FUNCTION "SEQUENCE_TRANSFER" : Void   // FC9, LAD
{ S7_Optimized_Access := 'TRUE' }
VERSION : 0.1
   VAR_TEMP   // added for the SCL form of the ladder/FBD networks
      _w1 : Bool;
      _w2 : Bool;
      _w3 : Bool;
      _w4 : Bool;
      _w5 : Bool;
      _w6 : Bool;
      _w7 : Bool;
      _w8 : Bool;
      _w9 : Bool;
      _w10 : Bool;
      _w11 : Bool;
      _w12 : Bool;
      _w13 : Bool;
      _w14 : Bool;
      _w15 : Bool;
      _w16 : Bool;
      _w17 : Bool;
      _w18 : Bool;
      _s5time1 : S5Time;
      _s5time2 : S5Time;
   END_VAR
BEGIN

REGION Network 1: START TRANSFER
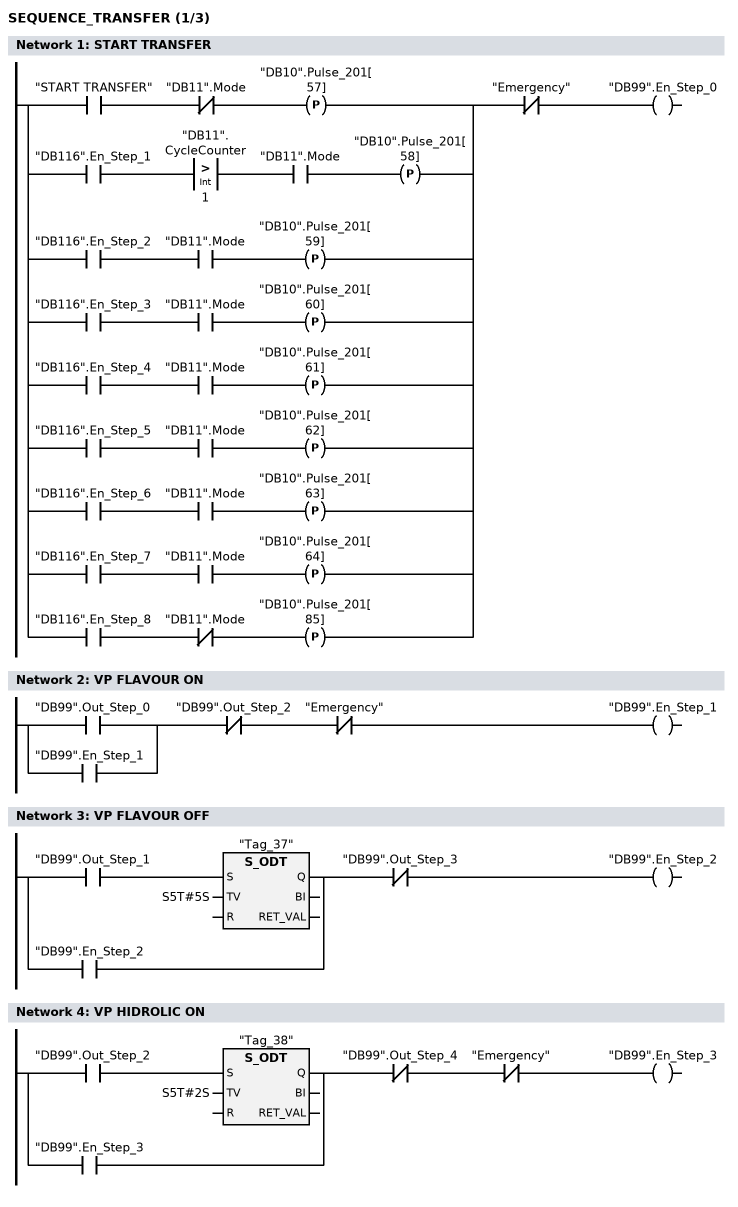
   RUNG wire#powerrail
      Contact( "START TRANSFER" )
      I_Contact( "DB11".Mode )
      P_Trig( "DB10".Pulse_201[57] )
      wire#w1
      I_Contact( "Emergency" )
      Coil( "DB99".En_Step_0 )
   END_RUNG
   RUNG wire#powerrail
      Contact( "DB116".En_Step_1 )
      { S7_Templates := "SrcType := Int" } GT_Contact(in1 := "DB11".CycleCounter, in2 := 1)
      Contact( "DB11".Mode )
      P_Trig( "DB10".Pulse_201[58] )
   END_RUNG wire#w1
   RUNG wire#powerrail
      Contact( "DB116".En_Step_2 )
      Contact( "DB11".Mode )
      P_Trig( "DB10".Pulse_201[59] )
   END_RUNG wire#w1
   RUNG wire#powerrail
      Contact( "DB116".En_Step_3 )
      Contact( "DB11".Mode )
      P_Trig( "DB10".Pulse_201[60] )
   END_RUNG wire#w1
   RUNG wire#powerrail
      Contact( "DB116".En_Step_4 )
      Contact( "DB11".Mode )
      P_Trig( "DB10".Pulse_201[61] )
   END_RUNG wire#w1
   RUNG wire#powerrail
      Contact( "DB116".En_Step_5 )
      Contact( "DB11".Mode )
      P_Trig( "DB10".Pulse_201[62] )
   END_RUNG wire#w1
   RUNG wire#powerrail
      Contact( "DB116".En_Step_6 )
      Contact( "DB11".Mode )
      P_Trig( "DB10".Pulse_201[63] )
   END_RUNG wire#w1
   RUNG wire#powerrail
      Contact( "DB116".En_Step_7 )
      Contact( "DB11".Mode )
      P_Trig( "DB10".Pulse_201[64] )
   END_RUNG wire#w1
   RUNG wire#powerrail
      Contact( "DB116".En_Step_8 )
      I_Contact( "DB11".Mode )
      P_Trig( "DB10".Pulse_201[85] )
   END_RUNG wire#w1
   // the same network as SCL:
   #_w1 := "START TRANSFER" AND NOT "DB11".Mode;
   #_w2 := #_w1 AND NOT "DB10".Pulse_201[57];   // rising edge
   "DB10".Pulse_201[57] := #_w1;
   #_w3 := "DB116".En_Step_1 AND ("DB11".CycleCounter > 1) AND "DB11".Mode;
   #_w4 := #_w3 AND NOT "DB10".Pulse_201[58];   // rising edge
   "DB10".Pulse_201[58] := #_w3;
   #_w5 := "DB116".En_Step_2 AND "DB11".Mode;
   #_w6 := #_w5 AND NOT "DB10".Pulse_201[59];   // rising edge
   "DB10".Pulse_201[59] := #_w5;
   #_w7 := "DB116".En_Step_3 AND "DB11".Mode;
   #_w8 := #_w7 AND NOT "DB10".Pulse_201[60];   // rising edge
   "DB10".Pulse_201[60] := #_w7;
   #_w9 := "DB116".En_Step_4 AND "DB11".Mode;
   #_w10 := #_w9 AND NOT "DB10".Pulse_201[61];   // rising edge
   "DB10".Pulse_201[61] := #_w9;
   #_w11 := "DB116".En_Step_5 AND "DB11".Mode;
   #_w12 := #_w11 AND NOT "DB10".Pulse_201[62];   // rising edge
   "DB10".Pulse_201[62] := #_w11;
   #_w13 := "DB116".En_Step_6 AND "DB11".Mode;
   #_w14 := #_w13 AND NOT "DB10".Pulse_201[63];   // rising edge
   "DB10".Pulse_201[63] := #_w13;
   #_w15 := "DB116".En_Step_7 AND "DB11".Mode;
   #_w16 := #_w15 AND NOT "DB10".Pulse_201[64];   // rising edge
   "DB10".Pulse_201[64] := #_w15;
   #_w17 := "DB116".En_Step_8 AND NOT "DB11".Mode;
   #_w18 := #_w17 AND NOT "DB10".Pulse_201[85];   // rising edge
   "DB10".Pulse_201[85] := #_w17;
   "DB99".En_Step_0 := (#_w2 OR #_w4 OR #_w6 OR #_w8 OR #_w10 OR #_w12 OR #_w14 OR #_w16 OR #_w18) AND NOT "Emergency";
END_REGION

REGION Network 2: VP FLAVOUR ON
   RUNG wire#powerrail
      Contact( "DB99".Out_Step_0 )
      wire#w1
      I_Contact( "DB99".Out_Step_2 )
      I_Contact( "Emergency" )
      Coil( "DB99".En_Step_1 )
   END_RUNG
   RUNG wire#powerrail
      Contact( "DB99".En_Step_1 )
   END_RUNG wire#w1
   // the same network as SCL:
   "DB99".En_Step_1 := ("DB99".Out_Step_0 OR "DB99".En_Step_1) AND NOT "DB99".Out_Step_2 AND NOT "Emergency";
END_REGION

REGION Network 3: VP FLAVOUR OFF
   RUNG wire#powerrail
      Contact( "DB99".Out_Step_1 )
      S_ODT(T_NO := "Tag_37", TV := S5T#5S, R :=, BI =>, RET_VAL =>)
      wire#w1
      I_Contact( "DB99".Out_Step_3 )
      Coil( "DB99".En_Step_2 )
   END_RUNG
   RUNG wire#powerrail
      Contact( "DB99".En_Step_2 )
   END_RUNG wire#w1
   // the same network as SCL:
   #_s5time1 := S_ODT(T_NO := "Tag_37", S := "DB99".Out_Step_1, TV := S5T#5S, Q => #_w1);
   "DB99".En_Step_2 := (#_w1 OR "DB99".En_Step_2) AND NOT "DB99".Out_Step_3;
END_REGION

REGION Network 4: VP HIDROLIC ON
   RUNG wire#powerrail
      Contact( "DB99".Out_Step_2 )
      S_ODT(T_NO := "Tag_38", TV := S5T#2S, R :=, BI =>, RET_VAL =>)
      wire#w1
      I_Contact( "DB99".Out_Step_4 )
      I_Contact( "Emergency" )
      Coil( "DB99".En_Step_3 )
   END_RUNG
   RUNG wire#powerrail
      Contact( "DB99".En_Step_3 )
   END_RUNG wire#w1
   // the same network as SCL:
   #_s5time1 := S_ODT(T_NO := "Tag_38", S := "DB99".Out_Step_2, TV := S5T#2S, Q => #_w1);
   "DB99".En_Step_3 := (#_w1 OR "DB99".En_Step_3) AND NOT "DB99".Out_Step_4 AND NOT "Emergency";
END_REGION

REGION Network 5
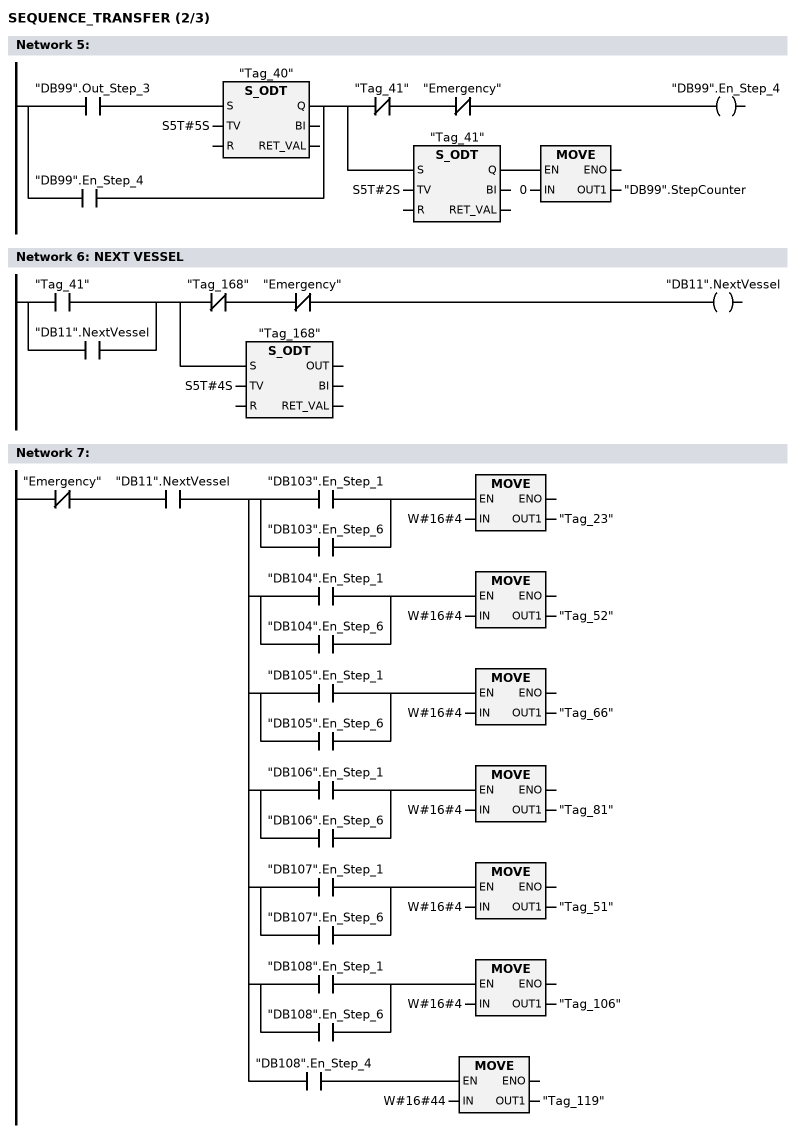
   RUNG wire#powerrail
      Contact( "DB99".Out_Step_3 )
      S_ODT(T_NO := "Tag_40", TV := S5T#5S, R :=, BI =>, RET_VAL =>)
      wire#w1
      I_Contact( "Tag_41" )
      I_Contact( "Emergency" )
      Coil( "DB99".En_Step_4 )
   END_RUNG
   RUNG wire#powerrail
      Contact( "DB99".En_Step_4 )
   END_RUNG wire#w1
   RUNG wire#w1
      S_ODT(T_NO := "Tag_41", TV := S5T#2S, R :=, BI =>, RET_VAL =>)
      Move(in := 0, out1 => "DB99".StepCounter)
   END_RUNG
   // the same network as SCL:
   #_s5time1 := S_ODT(T_NO := "Tag_40", S := "DB99".Out_Step_3, TV := S5T#5S, Q => #_w1);
   #_w2 := #_w1 OR "DB99".En_Step_4;
   "DB99".En_Step_4 := #_w2 AND NOT "Tag_41" AND NOT "Emergency";
   #_s5time2 := S_ODT(T_NO := "Tag_41", S := #_w2, TV := S5T#2S, Q => #_w3);
   IF #_w3 THEN "DB99".StepCounter := 0; END_IF;
END_REGION

REGION Network 6: NEXT VESSEL
   RUNG wire#powerrail
      Contact( "Tag_41" )
      wire#w1
      I_Contact( "Tag_168" )
      I_Contact( "Emergency" )
      Coil( "DB11".NextVessel )
   END_RUNG
   RUNG wire#powerrail
      Contact( "DB11".NextVessel )
   END_RUNG wire#w1
   RUNG wire#w1
      S_ODT(T_NO := "Tag_168", TV := S5T#4S, R :=, BI =>, RET_VAL =>)
   END_RUNG
   // the same network as SCL:
   #_w1 := "Tag_41" OR "DB11".NextVessel;
   "DB11".NextVessel := #_w1 AND NOT "Tag_168" AND NOT "Emergency";
   #_s5time1 := S_ODT(T_NO := "Tag_168", S := #_w1, TV := S5T#4S);
END_REGION

REGION Network 7
   RUNG wire#powerrail
      I_Contact( "Emergency" )
      Contact( "DB11".NextVessel )
      wire#w1
      Contact( "DB103".En_Step_1 )
      wire#w2
      Move(in := W#16#4, out1 => "Tag_23")
   END_RUNG
   RUNG wire#w1
      Contact( "DB103".En_Step_6 )
   END_RUNG wire#w2
   RUNG wire#w1
      Contact( "DB104".En_Step_1 )
      wire#w3
      Move(in := W#16#4, out1 => "Tag_52")
   END_RUNG
   RUNG wire#w1
      Contact( "DB104".En_Step_6 )
   END_RUNG wire#w3
   RUNG wire#w1
      Contact( "DB105".En_Step_1 )
      wire#w4
      Move(in := W#16#4, out1 => "Tag_66")
   END_RUNG
   RUNG wire#w1
      Contact( "DB105".En_Step_6 )
   END_RUNG wire#w4
   RUNG wire#w1
      Contact( "DB106".En_Step_1 )
      wire#w5
      Move(in := W#16#4, out1 => "Tag_81")
   END_RUNG
   RUNG wire#w1
      Contact( "DB106".En_Step_6 )
   END_RUNG wire#w5
   RUNG wire#w1
      Contact( "DB107".En_Step_1 )
      wire#w6
      Move(in := W#16#4, out1 => "Tag_51")
   END_RUNG
   RUNG wire#w1
      Contact( "DB107".En_Step_6 )
   END_RUNG wire#w6
   RUNG wire#w1
      Contact( "DB108".En_Step_1 )
      wire#w7
      Move(in := W#16#4, out1 => "Tag_106")
   END_RUNG
   RUNG wire#w1
      Contact( "DB108".En_Step_6 )
   END_RUNG wire#w7
   RUNG wire#w1
      Contact( "DB108".En_Step_4 )
      Move(in := W#16#44, out1 => "Tag_119")
   END_RUNG
   // the same network as SCL:
   #_w1 := NOT "Emergency" AND "DB11".NextVessel;
   IF #_w1 AND ("DB103".En_Step_1 OR "DB103".En_Step_6) THEN "Tag_23" := W#16#4; END_IF;
   IF #_w1 AND ("DB104".En_Step_1 OR "DB104".En_Step_6) THEN "Tag_52" := W#16#4; END_IF;
   IF #_w1 AND ("DB105".En_Step_1 OR "DB105".En_Step_6) THEN "Tag_66" := W#16#4; END_IF;
   IF #_w1 AND ("DB106".En_Step_1 OR "DB106".En_Step_6) THEN "Tag_81" := W#16#4; END_IF;
   IF #_w1 AND ("DB107".En_Step_1 OR "DB107".En_Step_6) THEN "Tag_51" := W#16#4; END_IF;
   IF #_w1 AND ("DB108".En_Step_1 OR "DB108".En_Step_6) THEN "Tag_106" := W#16#4; END_IF;
   IF #_w1 AND "DB108".En_Step_4 THEN "Tag_119" := W#16#44; END_IF;
END_REGION

REGION Network 8
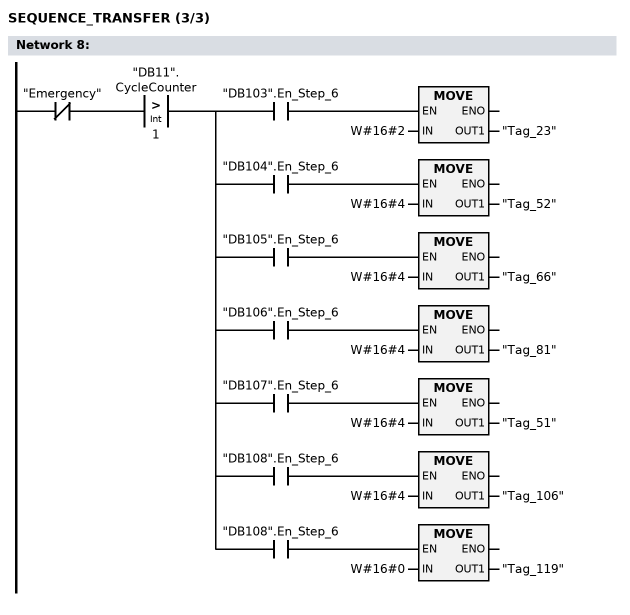
   RUNG wire#powerrail
      I_Contact( "Emergency" )
      { S7_Templates := "SrcType := Int" } GT_Contact(in1 := "DB11".CycleCounter, in2 := 1)
      wire#w1
      Contact( "DB103".En_Step_6 )
      Move(in := W#16#2, out1 => "Tag_23")
   END_RUNG
   RUNG wire#w1
      Contact( "DB104".En_Step_6 )
      Move(in := W#16#4, out1 => "Tag_52")
   END_RUNG
   RUNG wire#w1
      Contact( "DB105".En_Step_6 )
      Move(in := W#16#4, out1 => "Tag_66")
   END_RUNG
   RUNG wire#w1
      Contact( "DB106".En_Step_6 )
      Move(in := W#16#4, out1 => "Tag_81")
   END_RUNG
   RUNG wire#w1
      Contact( "DB107".En_Step_6 )
      Move(in := W#16#4, out1 => "Tag_51")
   END_RUNG
   RUNG wire#w1
      Contact( "DB108".En_Step_6 )
      Move(in := W#16#4, out1 => "Tag_106")
   END_RUNG
   RUNG wire#w1
      Contact( "DB108".En_Step_6 )
      Move(in := W#16#0, out1 => "Tag_119")
   END_RUNG
   // the same network as SCL:
   #_w1 := NOT "Emergency" AND ("DB11".CycleCounter > 1);
   IF #_w1 AND "DB103".En_Step_6 THEN "Tag_23" := W#16#2; END_IF;
   IF #_w1 AND "DB104".En_Step_6 THEN "Tag_52" := W#16#4; END_IF;
   IF #_w1 AND "DB105".En_Step_6 THEN "Tag_66" := W#16#4; END_IF;
   IF #_w1 AND "DB106".En_Step_6 THEN "Tag_81" := W#16#4; END_IF;
   IF #_w1 AND "DB107".En_Step_6 THEN "Tag_51" := W#16#4; END_IF;
   IF #_w1 AND "DB108".En_Step_6 THEN
       "Tag_106" := W#16#4;
       "Tag_119" := W#16#0;
   END_IF;
END_REGION
END_FUNCTION

FUNCTION "Cycle" : Void   // FC10, LAD
{ S7_Optimized_Access := 'TRUE' }
VERSION : 0.1
   VAR_TEMP   // added for the SCL form of the ladder/FBD networks
      _w1 : Bool;
      _w2 : Bool;
      _s5time1 : S5Time;
   END_VAR
BEGIN

REGION Network 1
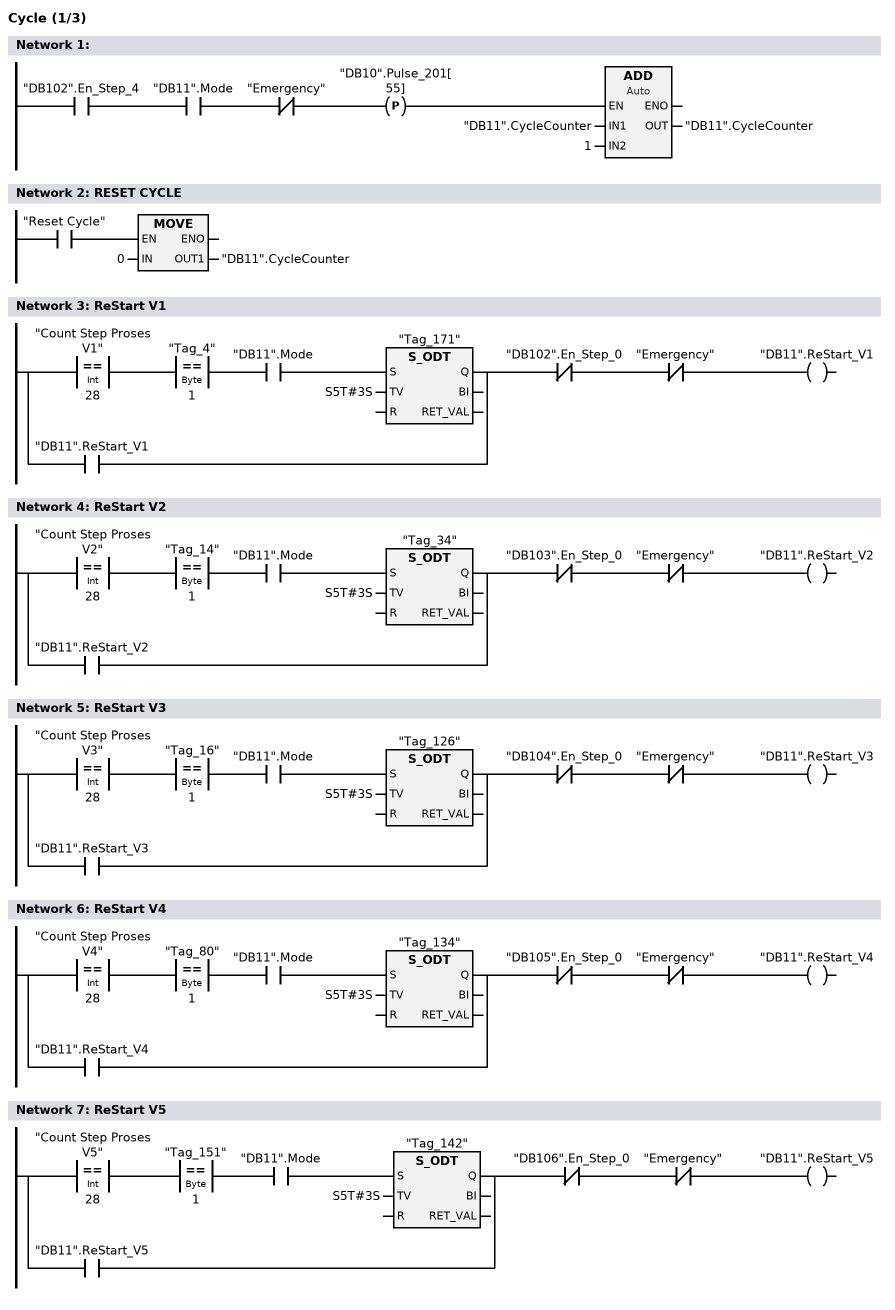
   RUNG wire#powerrail
      Contact( "DB102".En_Step_4 )
      Contact( "DB11".Mode )
      I_Contact( "Emergency" )
      P_Trig( "DB10".Pulse_201[55] )
      Add(in1 := "DB11".CycleCounter, in2 := 1, out => "DB11".CycleCounter)
   END_RUNG
   // the same network as SCL:
   #_w1 := "DB102".En_Step_4 AND "DB11".Mode AND NOT "Emergency";
   #_w2 := #_w1 AND NOT "DB10".Pulse_201[55];   // rising edge
   "DB10".Pulse_201[55] := #_w1;
   IF #_w2 THEN "DB11".CycleCounter := "DB11".CycleCounter + 1; END_IF;
END_REGION

REGION Network 2: RESET CYCLE
   RUNG wire#powerrail
      Contact( "Reset Cycle" )
      Move(in := 0, out1 => "DB11".CycleCounter)
   END_RUNG
   // the same network as SCL:
   IF "Reset Cycle" THEN "DB11".CycleCounter := 0; END_IF;
END_REGION

REGION Network 3: ReStart V1
   RUNG wire#powerrail
      { S7_Templates := "SrcType := Int" } EQ_Contact(in1 := "Count Step Proses V1", in2 := 28)
      { S7_Templates := "SrcType := Byte" } EQ_Contact(in1 := "Tag_4", in2 := 1)
      Contact( "DB11".Mode )
      S_ODT(T_NO := "Tag_171", TV := S5T#3S, R :=, BI =>, RET_VAL =>)
      wire#w1
      I_Contact( "DB102".En_Step_0 )
      I_Contact( "Emergency" )
      Coil( "DB11".ReStart_V1 )
   END_RUNG
   RUNG wire#powerrail
      Contact( "DB11".ReStart_V1 )
   END_RUNG wire#w1
   // the same network as SCL:
   #_s5time1 := S_ODT(T_NO := "Tag_171",
                      S := ("Count Step Proses V1" = 28) AND ("Tag_4" = 1) AND "DB11".Mode,
                      TV := S5T#3S,
                      Q => #_w1);
   "DB11".ReStart_V1 := (#_w1 OR "DB11".ReStart_V1) AND NOT "DB102".En_Step_0 AND NOT "Emergency";
END_REGION

REGION Network 4: ReStart V2
   RUNG wire#powerrail
      { S7_Templates := "SrcType := Int" } EQ_Contact(in1 := "Count Step Proses V2", in2 := 28)
      { S7_Templates := "SrcType := Byte" } EQ_Contact(in1 := "Tag_14", in2 := 1)
      Contact( "DB11".Mode )
      S_ODT(T_NO := "Tag_34", TV := S5T#3S, R :=, BI =>, RET_VAL =>)
      wire#w1
      I_Contact( "DB103".En_Step_0 )
      I_Contact( "Emergency" )
      Coil( "DB11".ReStart_V2 )
   END_RUNG
   RUNG wire#powerrail
      Contact( "DB11".ReStart_V2 )
   END_RUNG wire#w1
   // the same network as SCL:
   #_s5time1 := S_ODT(T_NO := "Tag_34",
                      S := ("Count Step Proses V2" = 28) AND ("Tag_14" = 1) AND "DB11".Mode,
                      TV := S5T#3S,
                      Q => #_w1);
   "DB11".ReStart_V2 := (#_w1 OR "DB11".ReStart_V2) AND NOT "DB103".En_Step_0 AND NOT "Emergency";
END_REGION

REGION Network 5: ReStart V3
   RUNG wire#powerrail
      { S7_Templates := "SrcType := Int" } EQ_Contact(in1 := "Count Step Proses V3", in2 := 28)
      { S7_Templates := "SrcType := Byte" } EQ_Contact(in1 := "Tag_16", in2 := 1)
      Contact( "DB11".Mode )
      S_ODT(T_NO := "Tag_126", TV := S5T#3S, R :=, BI =>, RET_VAL =>)
      wire#w1
      I_Contact( "DB104".En_Step_0 )
      I_Contact( "Emergency" )
      Coil( "DB11".ReStart_V3 )
   END_RUNG
   RUNG wire#powerrail
      Contact( "DB11".ReStart_V3 )
   END_RUNG wire#w1
   // the same network as SCL:
   #_s5time1 := S_ODT(T_NO := "Tag_126",
                      S := ("Count Step Proses V3" = 28) AND ("Tag_16" = 1) AND "DB11".Mode,
                      TV := S5T#3S,
                      Q => #_w1);
   "DB11".ReStart_V3 := (#_w1 OR "DB11".ReStart_V3) AND NOT "DB104".En_Step_0 AND NOT "Emergency";
END_REGION

REGION Network 6: ReStart V4
   RUNG wire#powerrail
      { S7_Templates := "SrcType := Int" } EQ_Contact(in1 := "Count Step Proses V4", in2 := 28)
      { S7_Templates := "SrcType := Byte" } EQ_Contact(in1 := "Tag_80", in2 := 1)
      Contact( "DB11".Mode )
      S_ODT(T_NO := "Tag_134", TV := S5T#3S, R :=, BI =>, RET_VAL =>)
      wire#w1
      I_Contact( "DB105".En_Step_0 )
      I_Contact( "Emergency" )
      Coil( "DB11".ReStart_V4 )
   END_RUNG
   RUNG wire#powerrail
      Contact( "DB11".ReStart_V4 )
   END_RUNG wire#w1
   // the same network as SCL:
   #_s5time1 := S_ODT(T_NO := "Tag_134",
                      S := ("Count Step Proses V4" = 28) AND ("Tag_80" = 1) AND "DB11".Mode,
                      TV := S5T#3S,
                      Q => #_w1);
   "DB11".ReStart_V4 := (#_w1 OR "DB11".ReStart_V4) AND NOT "DB105".En_Step_0 AND NOT "Emergency";
END_REGION

REGION Network 7: ReStart V5
   RUNG wire#powerrail
      { S7_Templates := "SrcType := Int" } EQ_Contact(in1 := "Count Step Proses V5", in2 := 28)
      { S7_Templates := "SrcType := Byte" } EQ_Contact(in1 := "Tag_151", in2 := 1)
      Contact( "DB11".Mode )
      S_ODT(T_NO := "Tag_142", TV := S5T#3S, R :=, BI =>, RET_VAL =>)
      wire#w1
      I_Contact( "DB106".En_Step_0 )
      I_Contact( "Emergency" )
      Coil( "DB11".ReStart_V5 )
   END_RUNG
   RUNG wire#powerrail
      Contact( "DB11".ReStart_V5 )
   END_RUNG wire#w1
   // the same network as SCL:
   #_s5time1 := S_ODT(T_NO := "Tag_142",
                      S := ("Count Step Proses V5" = 28) AND ("Tag_151" = 1) AND "DB11".Mode,
                      TV := S5T#3S,
                      Q => #_w1);
   "DB11".ReStart_V5 := (#_w1 OR "DB11".ReStart_V5) AND NOT "DB106".En_Step_0 AND NOT "Emergency";
END_REGION

REGION Network 8: ReStart V6
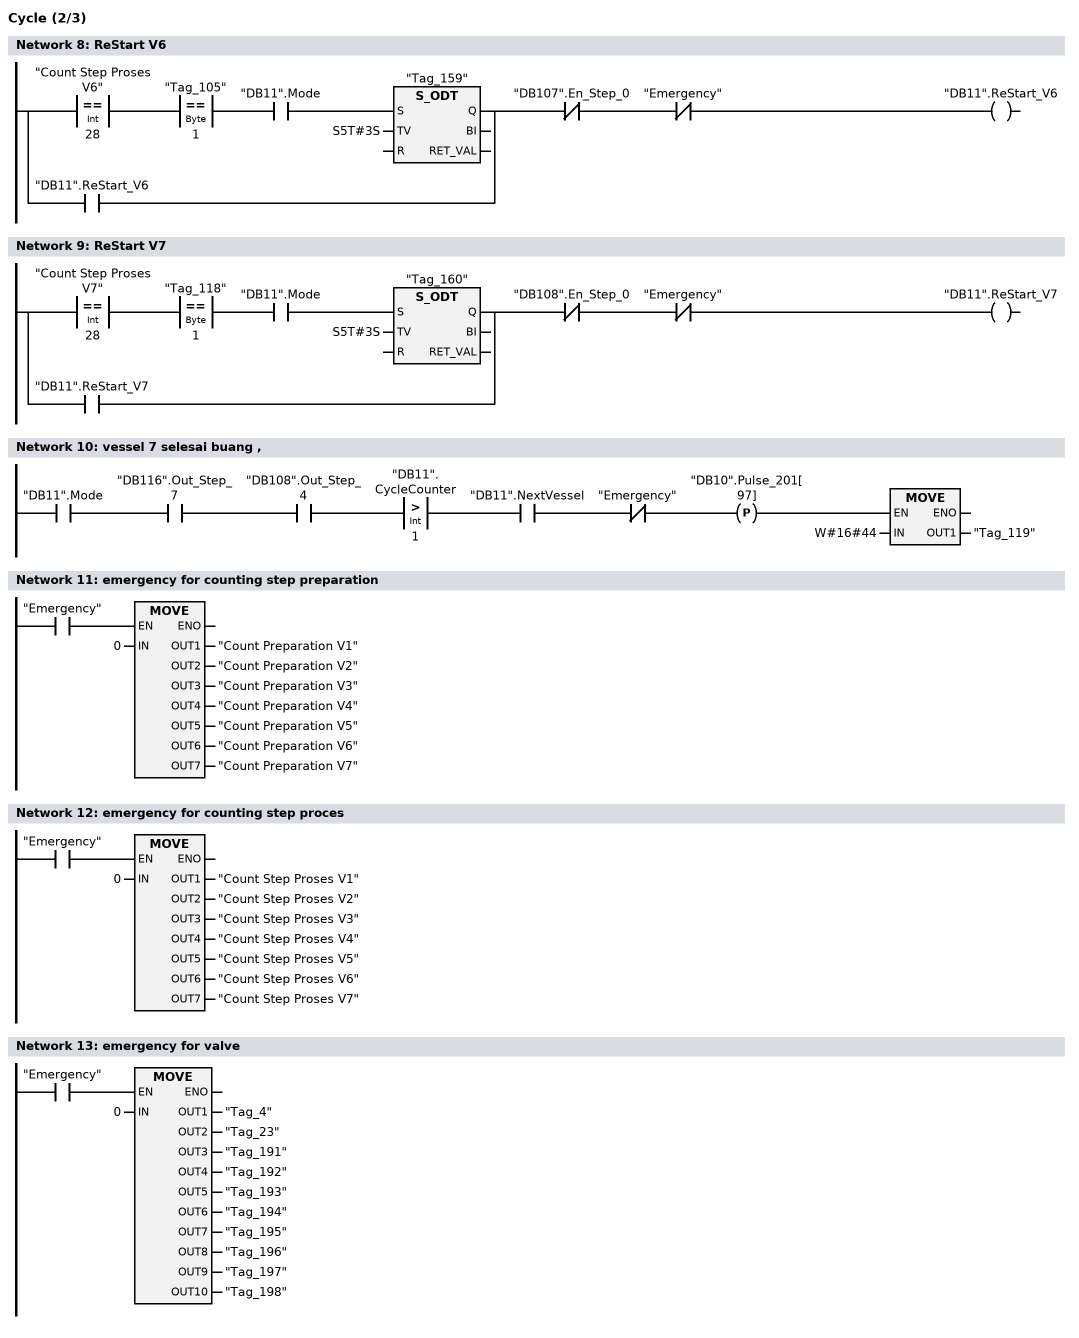
   RUNG wire#powerrail
      { S7_Templates := "SrcType := Int" } EQ_Contact(in1 := "Count Step Proses V6", in2 := 28)
      { S7_Templates := "SrcType := Byte" } EQ_Contact(in1 := "Tag_105", in2 := 1)
      Contact( "DB11".Mode )
      S_ODT(T_NO := "Tag_159", TV := S5T#3S, R :=, BI =>, RET_VAL =>)
      wire#w1
      I_Contact( "DB107".En_Step_0 )
      I_Contact( "Emergency" )
      Coil( "DB11".ReStart_V6 )
   END_RUNG
   RUNG wire#powerrail
      Contact( "DB11".ReStart_V6 )
   END_RUNG wire#w1
   // the same network as SCL:
   #_s5time1 := S_ODT(T_NO := "Tag_159",
                      S := ("Count Step Proses V6" = 28) AND ("Tag_105" = 1) AND "DB11".Mode,
                      TV := S5T#3S,
                      Q => #_w1);
   "DB11".ReStart_V6 := (#_w1 OR "DB11".ReStart_V6) AND NOT "DB107".En_Step_0 AND NOT "Emergency";
END_REGION

REGION Network 9: ReStart V7
   RUNG wire#powerrail
      { S7_Templates := "SrcType := Int" } EQ_Contact(in1 := "Count Step Proses V7", in2 := 28)
      { S7_Templates := "SrcType := Byte" } EQ_Contact(in1 := "Tag_118", in2 := 1)
      Contact( "DB11".Mode )
      S_ODT(T_NO := "Tag_160", TV := S5T#3S, R :=, BI =>, RET_VAL =>)
      wire#w1
      I_Contact( "DB108".En_Step_0 )
      I_Contact( "Emergency" )
      Coil( "DB11".ReStart_V7 )
   END_RUNG
   RUNG wire#powerrail
      Contact( "DB11".ReStart_V7 )
   END_RUNG wire#w1
   // the same network as SCL:
   #_s5time1 := S_ODT(T_NO := "Tag_160",
                      S := ("Count Step Proses V7" = 28) AND ("Tag_118" = 1) AND "DB11".Mode,
                      TV := S5T#3S,
                      Q => #_w1);
   "DB11".ReStart_V7 := (#_w1 OR "DB11".ReStart_V7) AND NOT "DB108".En_Step_0 AND NOT "Emergency";
END_REGION

REGION Network 10: vessel 7 selesai buang ,
   RUNG wire#powerrail
      Contact( "DB11".Mode )
      Contact( "DB116".Out_Step_7 )
      Contact( "DB108".Out_Step_4 )
      { S7_Templates := "SrcType := Int" } GT_Contact(in1 := "DB11".CycleCounter, in2 := 1)
      Contact( "DB11".NextVessel )
      I_Contact( "Emergency" )
      P_Trig( "DB10".Pulse_201[97] )
      Move(in := W#16#44, out1 => "Tag_119")
   END_RUNG
   // the same network as SCL:
   #_w1 := "DB11".Mode AND "DB116".Out_Step_7 AND "DB108".Out_Step_4 AND ("DB11".CycleCounter > 1) AND "DB11".NextVessel AND NOT "Emergency";
   #_w2 := #_w1 AND NOT "DB10".Pulse_201[97];   // rising edge
   "DB10".Pulse_201[97] := #_w1;
   IF #_w2 THEN "Tag_119" := W#16#44; END_IF;
END_REGION

REGION Network 11: emergency for counting step preparation
   RUNG wire#powerrail
      Contact( "Emergency" )
      Move(in := 0, out1 => "Count Preparation V1", out2 => "Count Preparation V2", out3 => "Count Preparation V3", out4 => "Count Preparation V4", out5 => "Count Preparation V5", out6 => "Count Preparation V6", out7 => "Count Preparation V7")
   END_RUNG
   // the same network as SCL:
   IF "Emergency" THEN
       "Count Preparation V1" := 0;
       "Count Preparation V2" := 0;
       "Count Preparation V3" := 0;
       "Count Preparation V4" := 0;
       "Count Preparation V5" := 0;
       "Count Preparation V6" := 0;
       "Count Preparation V7" := 0;
   END_IF;
END_REGION

REGION Network 12: emergency for counting step proces
   RUNG wire#powerrail
      Contact( "Emergency" )
      Move(in := 0, out1 => "Count Step Proses V1", out2 => "Count Step Proses V2", out3 => "Count Step Proses V3", out4 => "Count Step Proses V4", out5 => "Count Step Proses V5", out6 => "Count Step Proses V6", out7 => "Count Step Proses V7")
   END_RUNG
   // the same network as SCL:
   IF "Emergency" THEN
       "Count Step Proses V1" := 0;
       "Count Step Proses V2" := 0;
       "Count Step Proses V3" := 0;
       "Count Step Proses V4" := 0;
       "Count Step Proses V5" := 0;
       "Count Step Proses V6" := 0;
       "Count Step Proses V7" := 0;
   END_IF;
END_REGION

REGION Network 13: emergency for valve
   RUNG wire#powerrail
      Contact( "Emergency" )
      Move(in := 0, out1 => "Tag_4", out2 => "Tag_23", out3 => "Tag_191", out4 => "Tag_192", out5 => "Tag_193", out6 => "Tag_194", out7 => "Tag_195", out8 => "Tag_196", out9 => "Tag_197", out10 => "Tag_198")
   END_RUNG
   // the same network as SCL:
   IF "Emergency" THEN
       "Tag_4" := 0;
       "Tag_23" := 0;
       "Tag_191" := 0;
       "Tag_192" := 0;
       "Tag_193" := 0;
       "Tag_194" := 0;
       "Tag_195" := 0;
       "Tag_196" := 0;
       "Tag_197" := 0;
       "Tag_198" := 0;
   END_IF;
END_REGION

REGION Network 14: emergency
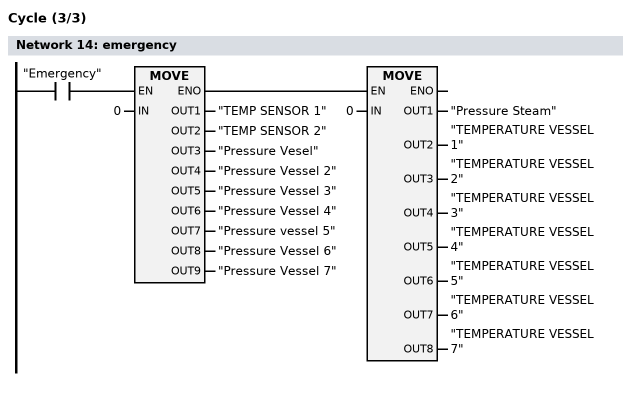
   RUNG wire#powerrail
      Contact( "Emergency" )
      Move(in := 0, out1 => "TEMP SENSOR 1", out2 => "TEMP SENSOR 2", out3 => "Pressure Vesel", out4 => "Pressure Vessel 2", out5 => "Pressure Vessel 3", out6 => "Pressure Vessel 4", out7 => "Pressure vessel 5", out8 => "Pressure Vessel 6", out9 => "Pressure Vessel 7")
      Move(in := 0, out1 => "Pressure Steam", out2 => "TEMPERATURE VESSEL 1", out3 => "TEMPERATURE VESSEL 2", out4 => "TEMPERATURE VESSEL 3", out5 => "TEMPERATURE VESSEL 4", out6 => "TEMPERATURE VESSEL 5", out7 => "TEMPERATURE VESSEL 6", out8 => "TEMPERATURE VESSEL 7")
   END_RUNG
   // the same network as SCL:
   IF "Emergency" THEN
       "TEMP SENSOR 1" := 0;
       "TEMP SENSOR 2" := 0;
       "Pressure Vesel" := 0;
       "Pressure Vessel 2" := 0;
       "Pressure Vessel 3" := 0;
       "Pressure Vessel 4" := 0;
       "Pressure vessel 5" := 0;
       "Pressure Vessel 6" := 0;
       "Pressure Vessel 7" := 0;
       "Pressure Steam" := 0;
       "TEMPERATURE VESSEL 1" := 0;
       "TEMPERATURE VESSEL 2" := 0;
       "TEMPERATURE VESSEL 3" := 0;
       "TEMPERATURE VESSEL 4" := 0;
       "TEMPERATURE VESSEL 5" := 0;
       "TEMPERATURE VESSEL 6" := 0;
       "TEMPERATURE VESSEL 7" := 0;
   END_IF;
END_REGION
END_FUNCTION

FUNCTION "VESSEL 2 PROSES" : Void   // FC11, LAD
{ S7_Optimized_Access := 'TRUE' }
VERSION : 0.1
   VAR_TEMP   // added for the SCL form of the ladder/FBD networks
      _w1 : Bool;
      _w2 : Bool;
   END_VAR
BEGIN

REGION Network 1: BUKA VALVE VP 12 DAN VP 17
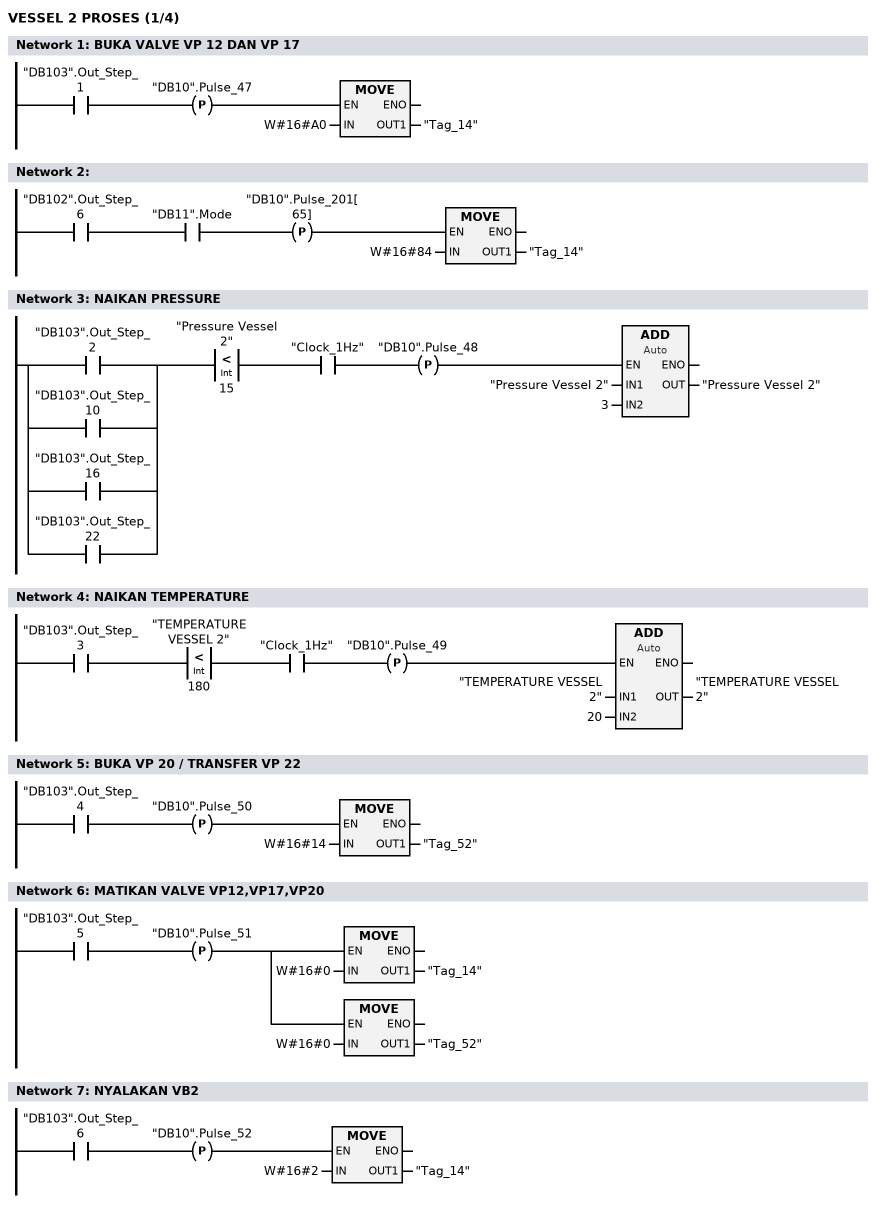
   RUNG wire#powerrail
      Contact( "DB103".Out_Step_1 )
      P_Trig( "DB10".Pulse_47 )
      Move(in := W#16#A0, out1 => "Tag_14")
   END_RUNG
   // the same network as SCL:
   #_w1 := "DB103".Out_Step_1 AND NOT "DB10".Pulse_47;   // rising edge
   "DB10".Pulse_47 := "DB103".Out_Step_1;
   IF #_w1 THEN "Tag_14" := W#16#A0; END_IF;
END_REGION

REGION Network 2
   RUNG wire#powerrail
      Contact( "DB102".Out_Step_6 )
      Contact( "DB11".Mode )
      P_Trig( "DB10".Pulse_201[65] )
      Move(in := W#16#84, out1 => "Tag_14")
   END_RUNG
   // the same network as SCL:
   #_w1 := "DB102".Out_Step_6 AND "DB11".Mode;
   #_w2 := #_w1 AND NOT "DB10".Pulse_201[65];   // rising edge
   "DB10".Pulse_201[65] := #_w1;
   IF #_w2 THEN "Tag_14" := W#16#84; END_IF;
END_REGION

REGION Network 3: NAIKAN PRESSURE
   RUNG wire#powerrail
      Contact( "DB103".Out_Step_2 )
      wire#w1
      { S7_Templates := "SrcType := Int" } LT_Contact(in1 := "Pressure Vessel 2", in2 := 15)
      Contact( "Clock_1Hz" )
      P_Trig( "DB10".Pulse_48 )
      Add(in1 := "Pressure Vessel 2", in2 := 3, out => "Pressure Vessel 2")
   END_RUNG
   RUNG wire#powerrail
      Contact( "DB103".Out_Step_10 )
   END_RUNG wire#w1
   RUNG wire#powerrail
      Contact( "DB103".Out_Step_16 )
   END_RUNG wire#w1
   RUNG wire#powerrail
      Contact( "DB103".Out_Step_22 )
   END_RUNG wire#w1
   // the same network as SCL:
   #_w1 := ("DB103".Out_Step_2 OR "DB103".Out_Step_10 OR "DB103".Out_Step_16 OR "DB103".Out_Step_22) AND ("Pressure Vessel 2" < 15) AND "Clock_1Hz";
   #_w2 := #_w1 AND NOT "DB10".Pulse_48;   // rising edge
   "DB10".Pulse_48 := #_w1;
   IF #_w2 THEN "Pressure Vessel 2" := "Pressure Vessel 2" + 3; END_IF;
END_REGION

REGION Network 4: NAIKAN TEMPERATURE
   RUNG wire#powerrail
      Contact( "DB103".Out_Step_3 )
      { S7_Templates := "SrcType := Int" } LT_Contact(in1 := "TEMPERATURE VESSEL 2", in2 := 180)
      Contact( "Clock_1Hz" )
      P_Trig( "DB10".Pulse_49 )
      Add(in1 := "TEMPERATURE VESSEL 2", in2 := 20, out => "TEMPERATURE VESSEL 2")
   END_RUNG
   // the same network as SCL:
   #_w1 := "DB103".Out_Step_3 AND ("TEMPERATURE VESSEL 2" < 180) AND "Clock_1Hz";
   #_w2 := #_w1 AND NOT "DB10".Pulse_49;   // rising edge
   "DB10".Pulse_49 := #_w1;
   IF #_w2 THEN "TEMPERATURE VESSEL 2" := "TEMPERATURE VESSEL 2" + 20; END_IF;
END_REGION

REGION Network 5: BUKA VP 20 / TRANSFER VP 22
   RUNG wire#powerrail
      Contact( "DB103".Out_Step_4 )
      P_Trig( "DB10".Pulse_50 )
      Move(in := W#16#14, out1 => "Tag_52")
   END_RUNG
   // the same network as SCL:
   #_w1 := "DB103".Out_Step_4 AND NOT "DB10".Pulse_50;   // rising edge
   "DB10".Pulse_50 := "DB103".Out_Step_4;
   IF #_w1 THEN "Tag_52" := W#16#14; END_IF;
END_REGION

REGION Network 6: MATIKAN VALVE VP12,VP17,VP20
   RUNG wire#powerrail
      Contact( "DB103".Out_Step_5 )
      P_Trig( "DB10".Pulse_51 )
      wire#w1
      Move(in := W#16#0, out1 => "Tag_14")
   END_RUNG
   RUNG wire#w1
      Move(in := W#16#0, out1 => "Tag_52")
   END_RUNG
   // the same network as SCL:
   #_w1 := "DB103".Out_Step_5 AND NOT "DB10".Pulse_51;   // rising edge
   "DB10".Pulse_51 := "DB103".Out_Step_5;
   IF #_w1 THEN
       "Tag_14" := W#16#0;
       "Tag_52" := W#16#0;
   END_IF;
END_REGION

REGION Network 7: NYALAKAN VB2
   RUNG wire#powerrail
      Contact( "DB103".Out_Step_6 )
      P_Trig( "DB10".Pulse_52 )
      Move(in := W#16#2, out1 => "Tag_14")
   END_RUNG
   // the same network as SCL:
   #_w1 := "DB103".Out_Step_6 AND NOT "DB10".Pulse_52;   // rising edge
   "DB10".Pulse_52 := "DB103".Out_Step_6;
   IF #_w1 THEN "Tag_14" := W#16#2; END_IF;
END_REGION

REGION Network 8: TURUNKAN PRESSURE